// TIA Portal project "Konzept_zur_Überwachung_der_Feuchtigkeit_des_Getriebeöls" (V18)

(* hardware
DEVICE "Haupt_Station"  TP2200 Comfort
   slot 0: "Haupt_Station"  TP2200 Comfort  6AV2 124-0XC02-0AX0  17.0.0.0
   slot 1: "HMI_RT"  TP2200 Comfort  6AV2 124-0XC02-0AX0  17.0.0.0
   slot 5: "Haupt_Station.IE_CP_2"  PROFINET Interface  17.0.0.0
      slot 1: "PROFINET Schnittstelle_1"  PROFINET Interface
         slot 1: "Port_1"  Port
         slot 2: "Port_2"  Port
   slot 6: "Haupt_Station.IE_CP_1"  PROFINET Interface  17.0.0.0
      slot 1: "PROFINET Schnittstelle_GBit"  PROFINET Interface
         slot 1: "Port_1"  Port
   slot 7: "Haupt_Station.MPI/DP_CP_1"  MPI/DP Interface  17.0.0.0
DEVICE "S7-1500/ET200MP-Station_1"  S7-1500 station
   slot 0: "Profilschiene_0"  Rack  6ES7 590-1***0-0AA0
   slot 1: "1513"  CPU 1513-1 PN  6ES7 513-1AM03-0AB0  V3.0
      slot 3: "CPU-Display_1"  6ES7591-1AA00-0AA0
      slot 32768: "PROFINET-Schnittstelle_1"  X1
         slot 32769: "Port_1"  X1 P1
         slot 32770: "Port_2"  X1 P2
      slot 34817: "Virtual CP interface port_1"  Virtual CP interface port  Virtual CP interface port
   slot 2: "DI 16x24VDC / DQ 16x24VDC/0.5A BA_1"  DI 16x24VDC/DQ 16x24VDC/0.5A BA  6ES7 523-1BL00-0AA0  V1.1
   slot 3: "AI 8xU/I/R/RTD BA_1"  AI 8xU/I/R/RTD BA  6ES7 531-7QF00-0AB0  V1.0
DEVICE "S7-300/ET200M-Station_1"  S7-300 station
   slot 0: "Profilschiene_0"  Rail  6ES7 390-1***0-0AA0
   slot 1: "PS 307 10A_1"  PS 307 10A  6ES7 307-1KA02-0AA0
   slot 2: "313C"  CPU 313C-2 DP  6ES7 313-6CG04-0AB0  V3.3
      slot 0: "MPI-Schnittstelle_1"  MPI
      slot 1: "DP-Schnittstelle_1"  DP
      slot 2: "DI 16/DO 16_1"  DI16/DO16
      slot 4: "Zählen_1"  Counter
   slot 4: "AI 8x13BIT_1"  AI8x13Bit  6ES7 331-1KF02-0AB0
*)

// ===== PLC "1513"  CPU 1513-1 PN =====

VAR_GLOBAL   // PLC tag table "Standard-Variablentabelle"
   "LDH_Temp_1(1)" AT %IW34 : Int;
   "LDH_Feucht_1(1)" AT %IW36 : Int;
   "LDH_Temp_2(1)" AT %IW38 : Int;
   "LDH_Feucht_2(1)" AT %IW40 : Int;
   "Gill_Fine(1)" AT %IW42 : Int;
   "Gill_Coarse(1)" AT %IW44 : Int;
   "Gill_Water(1)" AT %IW46 : Int;
   "Gill_Fehler(1)" AT %IW48 : Int;
   "Rote_Lampe(1)" AT %Q0.0 : Bool;
   "Orange_Lampe(1)" AT %Q0.1 : Bool;
   "Grüne_Lampe_2(1)" AT %Q0.2 : Bool;
   "Abschalten_M(1)" AT %Q0.3 : Bool;
   "Quittierung(1)" AT %I0.0 : Bool;
END_VAR

DATA_BLOCK "Rt_Zyklus_DB"   // DB1
{ S7_Optimized_Access := 'TRUE' }
VERSION : 0.1
// stored: InstanceOfName Rt_Zyklus
"Rt_Zyklus"
BEGIN
END_DATA_BLOCK

DATA_BLOCK "LDH100_DB_1"   // DB2
{ S7_Optimized_Access := 'TRUE' }
VERSION : 0.1
// stored: InstanceOfName LDH100
"LDH100"
BEGIN
END_DATA_BLOCK

DATA_BLOCK "LDH100_DB_2"   // DB3
{ S7_Optimized_Access := 'TRUE' }
VERSION : 0.1
// stored: InstanceOfName LDH100
"LDH100"
BEGIN
END_DATA_BLOCK

DATA_BLOCK "GILL4212_DB"   // DB4
{ S7_Optimized_Access := 'TRUE' }
VERSION : 0.1
// stored: InstanceOfName GILL4212
"GILL4212"
BEGIN
END_DATA_BLOCK

DATA_BLOCK "HMI"   // DB5
{ S7_Optimized_Access := 'TRUE' }
VERSION : 0.1
   VAR
      Quittieren1500 : Bool;
   END_VAR
BEGIN
END_DATA_BLOCK

FUNCTION_BLOCK "LDH100"   // FB1, SCL
{ S7_Optimized_Access := 'TRUE' }
VERSION : 0.1
   VAR_INPUT
      AI_Temp_RAW : Int;
      cycleTime_ms : Real;
      AI_Hum_RAW : Int;
      Quittieren : Bool;
   END_VAR
   VAR_OUTPUT
      Temp_filt : Real;
      Temp_real : Real;
      Hum_filt : Real;
      Hum_real : Real;
      Warnung : Bool;
      Alarm_Temp : Bool;
      Alarm_Hum : Bool;
      OK : Bool;
      SensorError_Temp : Bool;
      SensorError_Hum : Bool;
      SensorDefekt : Bool;
      Strom_Temp_mA : Real;
      Strom_Hum_mA : Real;
   END_VAR
   VAR
      Alarm_Temp_Intern : Bool;
      TempGrenze_Alarm : Real := 0.0;
      HumGrenze_Alarm : Real := 0.0;
      Alarm_Hum_Intern : Bool;
      intervall_temp : Real;
      intervall_hum : Real;
      TON_temp : TON_TIME;
      TON_Hum : TON_TIME;
      RawTol : Int;
      RawMin : Int;
      RawMax : Int;
   END_VAR
   VAR_TEMP
      Norm_Temp : Real;
      alpha_pt1 : Real;
      Norm_Hum : Real;
   END_VAR
   VAR CONSTANT
      T_PT1_ms : Real := 565.0;
   END_VAR
BEGIN
   // -2) Rohwert-Toleranz (±0,2 mA auf 4–>20 mA = -346–>27648)
   #RawTol := REAL_TO_INT((0.2 / 16.0) * 27648.0);
   #RawMin := - #RawTol;
   #RawMax := 27648 + #RawTol;

   // -1) Strom in mA berechnen
   #Strom_Temp_mA := (INT_TO_REAL(#AI_Temp_RAW) / 27648.0) * 16.0 + 4.0;
   #Strom_Hum_mA := (INT_TO_REAL(#AI_Hum_RAW) / 27648.0) * 16.0 + 4.0;

   // 0) Sensor-Error prüfen auf Rohwerte
   #SensorError_Temp := (#AI_Temp_RAW < #RawMin) OR (#AI_Temp_RAW > #RawMax);
   #SensorError_Hum := (#AI_Hum_RAW < #RawMin) OR (#AI_Hum_RAW > #RawMax);

   // 1) Skalierung in reale Werte
   #Temp_real := (INT_TO_REAL(#AI_Temp_RAW) / 27648.0) * 140.0 - 20.0;  // -20°C ... +120°C
   #Hum_real := (INT_TO_REAL(#AI_Hum_RAW) / 27648.0) * 100.0;         // 0% ... 100%

   // 2) Filter-Koeffizient berechnen (für τ = 565 ms → 90 % nach 1.3 s)
   #alpha_pt1 := #cycleTime_ms / (#T_PT1_ms + #cycleTime_ms);

   // 3) PT1-Glättung
   #Temp_filt := #Temp_filt + #alpha_pt1 * (#Temp_real - #Temp_filt);
   #Hum_filt := #Hum_filt + #alpha_pt1 * (#Hum_real - #Hum_filt);

   // 4) Alarm-Logik mit IEC-Timer (TON)
   // → nur auslösen, wenn Filterwert 1.3 s lang über Grenzwert liegt
   #TON_temp(IN := (#Temp_filt >= #TempGrenze_Alarm),
             PT := T#1300ms);
   #TON_Hum(IN := (#Hum_filt >= #HumGrenze_Alarm),
            PT := T#1300ms);

   IF #TON_temp.Q THEN
       #Alarm_Temp := TRUE;
   ELSIF #Quittieren AND (#Temp_filt < #TempGrenze_Alarm) THEN
       #Alarm_Temp := FALSE;
   END_IF;

   IF #TON_Hum.Q THEN
       #Alarm_Hum := TRUE;
   ELSIF #Quittieren AND (#Hum_filt < #HumGrenze_Alarm) THEN
       #Alarm_Hum := FALSE;
   END_IF;

   // 5) Warnung (Echtwerte, keine Filterung nötig)
   #Warnung := (#Temp_real >= (#TempGrenze_Alarm - #intervall_temp)) OR
   (#Hum_real >= (#HumGrenze_Alarm - #intervall_hum));

   // 6) OK-Status
   #OK := NOT #Alarm_Temp AND NOT #Alarm_Hum;
END_FUNCTION_BLOCK

FUNCTION_BLOCK "GILL4212"   // FB2, SCL
{ S7_Optimized_Access := 'TRUE' }
VERSION : 0.1
   VAR_INPUT
      AI_Fine_RAW : Int;
      AI_Coarse_RAW : Int;
      AI_Water_RAW : Int;
      Quittieren : Bool;
   END_VAR
   VAR_OUTPUT
      SensorError_Coarse : Bool;
      SensorError_Water : Bool;
      SensorError_Fine : Bool;
      Fine_percent : Real;
      Coarse_percent : Real;
      Water_percent : Real;
      Alarm_Wear : Bool;
      Alarm_Water : Bool;
      Warnung : Bool;
      OK : Bool;
   END_VAR
   VAR
      TON_Wear : TON_TIME;
      TON_Water : TON_TIME;
      Alarm_Wear_Intern : Bool;
      Alarm_Water_Intern : Bool;
      RawTol : Int;
      RawMin : Int;
      RawMax : Int;
   END_VAR
   VAR CONSTANT
      Wear_Alarm_Limit : Real := 70.0;
      Water_Alarm_Limit : Real := 60.0;
   END_VAR
BEGIN
   // -1) Toleranzbereich in Rohwert berechnen (±0.2 mA)
   #RawTol := REAL_TO_INT((0.2 / 16.0) * 27648.0);
   #RawMin := - #RawTol;
   #RawMax := 27648 + #RawTol;

   // 0) Rohwert auf Gültigkeit prüfen (Toleranz)
   #SensorError_Fine := (#AI_Fine_RAW < #RawMin) OR (#AI_Fine_RAW > #RawMax);
   #SensorError_Coarse := (#AI_Coarse_RAW < #RawMin) OR (#AI_Coarse_RAW > #RawMax);
   #SensorError_Water := (#AI_Water_RAW < #RawMin) OR (#AI_Water_RAW > #RawMax);

   // 1) Skalierung 4–20 mA → 0–100 %
   #Fine_percent := (INT_TO_REAL(#AI_Fine_RAW) / 27648.0) * 100.0;
   #Coarse_percent := (INT_TO_REAL(#AI_Coarse_RAW) / 27648.0) * 100.0;
   #Water_percent := (INT_TO_REAL(#AI_Water_RAW) / 27648.0) * 100.0;

   // 2) Alarmverzögerung (1,3 Sekunden) mit TON
   #TON_Wear(IN := (#Fine_percent >= #Wear_Alarm_Limit) OR (#Coarse_percent >= #Wear_Alarm_Limit), PT := T#1300ms);
   #TON_Water(IN := (#Water_percent >= #Water_Alarm_Limit), PT := T#1300ms);

   // 3) Alarm setzen nach Ablauf der Verzögerung
   IF #TON_Wear.Q THEN
       #Alarm_Wear_Intern := TRUE;
   END_IF;
   IF #TON_Water.Q THEN
       #Alarm_Water_Intern := TRUE;
   END_IF;

   // 4) Quittierung (nur wenn alle Werte unterhalb der Limits)
   IF #Quittieren AND #Fine_percent < #Wear_Alarm_Limit AND #Coarse_percent < #Wear_Alarm_Limit THEN
       #Alarm_Wear_Intern := FALSE;
   END_IF;
   IF #Quittieren AND #Water_percent < #Water_Alarm_Limit THEN
       #Alarm_Water_Intern := FALSE;
   END_IF;

   // 5) Ausgänge setzen
   #Alarm_Wear := #Alarm_Wear_Intern;
   #Alarm_Water := #Alarm_Water_Intern;

   // 6) Warnung (Vorwarnbereich ohne Verzögerung)
   #Warnung :=
   (#Fine_percent >= #Wear_Alarm_Limit - 20.0) OR
   (#Coarse_percent >= #Wear_Alarm_Limit - 20.0) OR
   (#Water_percent >= #Water_Alarm_Limit - 20.0);

   // 7) OK-Status
   #OK := NOT #Alarm_Wear AND NOT #Alarm_Water;
END_FUNCTION_BLOCK

FUNCTION_BLOCK "Rt_Zyklus"   // FB3, SCL
{ S7_Optimized_Access := 'TRUE' }
VERSION : 0.1
   VAR_INPUT
      Enable : Bool := True;
      Reset : Bool;
   END_VAR
   VAR_OUTPUT
      Cycle_ms : LReal;
      Min_ms : LReal;
      Max_ms : LReal;
      Error : Bool;
      Status : Int;
   END_VAR
   VAR
      Last_ns : LTime;
      Min_ns : LTime;
      Max_ns : LTime;
      ResetOld : Bool;
   END_VAR
BEGIN

   IF #Enable THEN

       // --- 1) Letzte Zykluszeit holen -----------------------------
       #Status := RT_INFO(
                          MODE := 25,          // MODE 25 = letzte Zykluszeit
                          OB := 0,
                          INFO := #Last_ns     // LTIME (Nanosekunden)
       );

   // Fehlerbehandlung -------------------------------------------
   #Error:= (#Status <> 0); // 0 = OK, alles andere = Fehler


       IF NOT #Error THEN

           // --- 2) Umrechnen in Millisekunden ----------------------
           #Cycle_ms := LINT_TO_LREAL(#Last_ns) / 1_000_000.0;

           // --- 3) Min/Max bilden ---------------------------------
           IF #Last_ns < #Min_ns THEN
               #Min_ns := #Last_ns;
           END_IF;

           IF #Last_ns > #Max_ns THEN
               #Max_ns := #Last_ns;
           END_IF;

           // --- 4) Reset per Flanke --------------------------------
           IF #Reset AND NOT #ResetOld THEN      // positive Flanke
               #Min_ns := #Last_ns;
               #Max_ns := #Last_ns;
           END_IF;

           // --- 5) Ausgänge aktualisieren --------------------------
           #Min_ms := LINT_TO_LREAL(#Min_ns) / 1_000_000.0;
           #Max_ms := LINT_TO_LREAL(#Max_ns) / 1_000_000.0;
       END_IF;

       // Flankenerkennung speicher­n
       #ResetOld := #Reset;

   ELSE
       // Messung deaktiviert → keine neuen Werte bilden
       #Error := FALSE;
       #Status := 0;
   END_IF;
END_FUNCTION_BLOCK

FUNCTION "Ampel_Logik" : Void   // FC1, SCL
{ S7_Optimized_Access := 'TRUE' }
VERSION : 0.1
   VAR_INPUT
      LDH1_Alarm_Hum : Bool;   // Alarm von LDH1 (Feuchte)
      LDH1_Alarm_Temp : Bool;   // Alarm von LDH1 (Temperatur)
      LDH2_Alarm_Hum : Bool;   // Alarm von LDH2 (Feuchte)
      LDH2_Alarm_Temp : Bool;   // Alarm von LDH2 (Temperatur)
      GILL_Alarm_Wear : Bool;   // Alarm vom GILL-Sensor (Verschleiß)
      GILL_Alarm_Water : Bool;   // Alarm vom GILL-Sensor (Wasser)
      LDH1_Warnung : Bool;   // Warnung LDH100_1
      LDH2_Warnung : Bool;   // Warnung LDH100_1
      GILL_Warnung : Bool;   // Warnung Verschleiss
   END_VAR
   VAR_OUTPUT
      LAMP_ROT : Bool;
      LAMP_ORANGE : Bool;
      LAMP_GRUEN : Bool;
   END_VAR
   VAR CONSTANT
      TempWarnMin : Real := 80.0;
      HumWarnMin : Real := 40.0;
      WearWarnMin : Real := 70.0;
      WaterWarnMin : Real := 50.0;
      HumAlarmLimit : Real := 100.0;
      TempAlarmLimit : Real := 60.0;
      WearAlarmLimit : Real := 80.0;
      WaterAlarmLimit : Real := 60.0;
   END_VAR
BEGIN
   // 1) ROT: mindestens ein Alarm-Flag aktiv
   IF #LDH1_Alarm_Hum OR #LDH1_Alarm_Temp OR
       #LDH2_Alarm_Hum OR #LDH2_Alarm_Temp OR
       #GILL_Alarm_Wear OR #GILL_Alarm_Water THEN

       #LAMP_ROT := TRUE;
       #LAMP_ORANGE := FALSE;
       #LAMP_GRUEN := FALSE;

       // 2) ORANGE: mindestens ein Wert im Warnbereich
       // 2) ORANGE: mindestens ein Warn-Flag aktiv
   ELSIF #LDH1_Warnung OR #LDH2_Warnung OR #GILL_Warnung THEN

       #LAMP_ROT := FALSE;
       #LAMP_ORANGE := TRUE;
       #LAMP_GRUEN := FALSE;

       // 3) GRÜN: alle Werte unter Warnschwelle
   ELSE
       #LAMP_ROT := FALSE;
       #LAMP_ORANGE := FALSE;
       #LAMP_GRUEN := TRUE;
   END_IF;
END_FUNCTION

ORGANIZATION_BLOCK "Main"   // OB1, LAD, ProgramCycle
TITLE = "Main Program Sweep (Cycle)"
{ S7_Optimized_Access := 'TRUE' }
VERSION : 0.1
   VAR_INPUT
      Initial_Call : Bool;   // Initial call of this OB
      Remanence : Bool;   // =True, if remanent data are available
   END_VAR
BEGIN

REGION Network 1
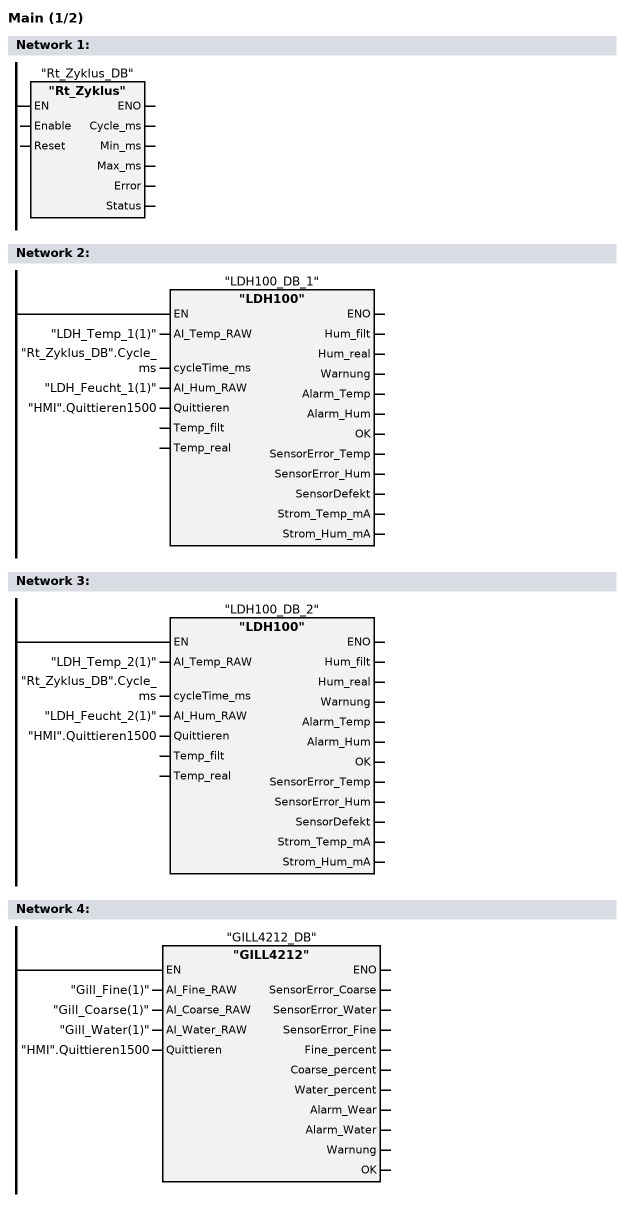
   RUNG wire#powerrail
      "Rt_Zyklus_DB"(Enable :=, Reset :=, Cycle_ms =>, Min_ms =>, Max_ms =>, Error =>, Status =>)
   END_RUNG
   // the same network as SCL:
   "Rt_Zyklus_DB"();   // "Rt_Zyklus"
END_REGION

REGION Network 2
   RUNG wire#powerrail
      "LDH100_DB_1"(AI_Temp_RAW := "LDH_Temp_1(1)", cycleTime_ms := "Rt_Zyklus_DB".Cycle_ms, AI_Hum_RAW := "LDH_Feucht_1(1)", Quittieren := "HMI".Quittieren1500, Temp_filt :=, Temp_real :=, Hum_filt =>, Hum_real =>, Warnung =>, Alarm_Temp =>, Alarm_Hum =>, OK =>, SensorError_Temp =>, SensorError_Hum =>, SensorDefekt =>, Strom_Temp_mA =>, Strom_Hum_mA =>)
   END_RUNG
   // the same network as SCL:
   "LDH100_DB_1"(AI_Temp_RAW := "LDH_Temp_1(1)",   // "LDH100"
                 cycleTime_ms := "Rt_Zyklus_DB".Cycle_ms,
                 AI_Hum_RAW := "LDH_Feucht_1(1)",
                 Quittieren := "HMI".Quittieren1500);
END_REGION

REGION Network 3
   RUNG wire#powerrail
      "LDH100_DB_2"(AI_Temp_RAW := "LDH_Temp_2(1)", cycleTime_ms := "Rt_Zyklus_DB".Cycle_ms, AI_Hum_RAW := "LDH_Feucht_2(1)", Quittieren := "HMI".Quittieren1500, Temp_filt :=, Temp_real :=, Hum_filt =>, Hum_real =>, Warnung =>, Alarm_Temp =>, Alarm_Hum =>, OK =>, SensorError_Temp =>, SensorError_Hum =>, SensorDefekt =>, Strom_Temp_mA =>, Strom_Hum_mA =>)
   END_RUNG
   // the same network as SCL:
   "LDH100_DB_2"(AI_Temp_RAW := "LDH_Temp_2(1)",   // "LDH100"
                 cycleTime_ms := "Rt_Zyklus_DB".Cycle_ms,
                 AI_Hum_RAW := "LDH_Feucht_2(1)",
                 Quittieren := "HMI".Quittieren1500);
END_REGION

REGION Network 4
   RUNG wire#powerrail
      "GILL4212_DB"(AI_Fine_RAW := "Gill_Fine(1)", AI_Coarse_RAW := "Gill_Coarse(1)", AI_Water_RAW := "Gill_Water(1)", Quittieren := "HMI".Quittieren1500, SensorError_Coarse =>, SensorError_Water =>, SensorError_Fine =>, Fine_percent =>, Coarse_percent =>, Water_percent =>, Alarm_Wear =>, Alarm_Water =>, Warnung =>, OK =>)
   END_RUNG
   // the same network as SCL:
   "GILL4212_DB"(AI_Fine_RAW := "Gill_Fine(1)",   // "GILL4212"
                 AI_Coarse_RAW := "Gill_Coarse(1)",
                 AI_Water_RAW := "Gill_Water(1)",
                 Quittieren := "HMI".Quittieren1500);
END_REGION

REGION Network 5
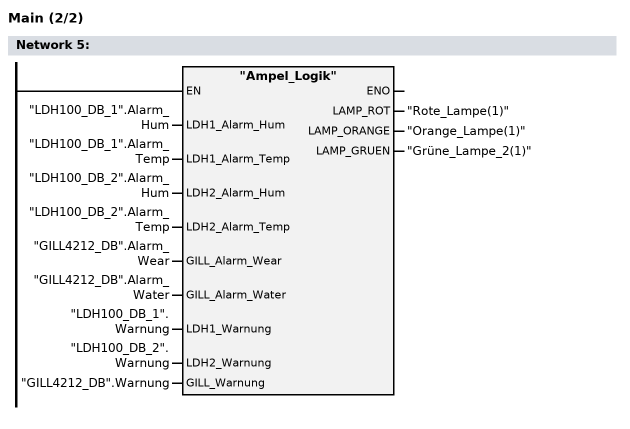
   RUNG wire#powerrail
      "Ampel_Logik"(LDH1_Alarm_Hum := "LDH100_DB_1".Alarm_Hum, LDH1_Alarm_Temp := "LDH100_DB_1".Alarm_Temp, LDH2_Alarm_Hum := "LDH100_DB_2".Alarm_Hum, LDH2_Alarm_Temp := "LDH100_DB_2".Alarm_Temp, GILL_Alarm_Wear := "GILL4212_DB".Alarm_Wear, GILL_Alarm_Water := "GILL4212_DB".Alarm_Water, LDH1_Warnung := "LDH100_DB_1".Warnung, LDH2_Warnung := "LDH100_DB_2".Warnung, GILL_Warnung := "GILL4212_DB".Warnung, LAMP_ROT => "Rote_Lampe(1)", LAMP_ORANGE => "Orange_Lampe(1)", LAMP_GRUEN => "Grüne_Lampe_2(1)")
   END_RUNG
   // the same network as SCL:
   "Ampel_Logik"(LDH1_Alarm_Hum := "LDH100_DB_1".Alarm_Hum,
                 LDH1_Alarm_Temp := "LDH100_DB_1".Alarm_Temp,
                 LDH2_Alarm_Hum := "LDH100_DB_2".Alarm_Hum,
                 LDH2_Alarm_Temp := "LDH100_DB_2".Alarm_Temp,
                 GILL_Alarm_Wear := "GILL4212_DB".Alarm_Wear,
                 GILL_Alarm_Water := "GILL4212_DB".Alarm_Water,
                 LDH1_Warnung := "LDH100_DB_1".Warnung,
                 LDH2_Warnung := "LDH100_DB_2".Warnung,
                 GILL_Warnung := "GILL4212_DB".Warnung,
                 LAMP_ROT => "Rote_Lampe(1)",
                 LAMP_ORANGE => "Orange_Lampe(1)",
                 LAMP_GRUEN => "Grüne_Lampe_2(1)");
END_REGION
END_ORGANIZATION_BLOCK

// ===== PLC "313C"  CPU 313C-2 DP =====

VAR_GLOBAL   // PLC tag table "Standard-Variablentabelle"
   "LDH_Temp_1" AT %IW272 : Int;
   "LDH_Feucht_1" AT %IW274 : Int;
   "LDH_Temp_2" AT %IW276 : Int;
   "LDH_Feucht_2" AT %IW278 : Int;
   "Gill_Fine" AT %IW280 : Int;
   "Gill_Coarse" AT %IW282 : Int;
   "Gill_Water" AT %IW284 : Int;
   "Gill_Fehler" AT %IW286 : Int;
   "Rote_Lampe" AT %I124.0 : Bool;
   "Orange_Lampe" AT %I124.1 : Bool;
   "Grüne_Lampe_2" AT %I124.2 : Bool;
   "Abschalten_M" AT %I124.3 : Bool;
END_VAR

VAR_GLOBAL   // PLC tag table "Merker_B"
   "B1" AT %M0.0 : Bool;
   "B2" AT %M0.1 : Bool;
   "B3" AT %M0.2 : Bool;
   "B4" AT %M0.3 : Bool;
   "B5" AT %M0.4 : Bool;
   "Re1" AT %MD1 : Real;
   "Re2" AT %MD2 : Real;
   "Re3" AT %MD3 : Real;
   "Re4" AT %MD4 : Real;
   "B7" AT %M0.6 : Bool;
   "B6" AT %M0.5 : Bool;
   "Re5" AT %MD5 : Real;
   "Re6" AT %MD6 : Real;
END_VAR

DATA_BLOCK "LDH100_DB_1"   // DB1
{ S7_Optimized_Access := 'FALSE' }
VERSION : 0.1
// stored: InstanceOfName LDH100
"LDH100"
BEGIN
   TempGrenze_Alarm := 60.0;
   HumGrenze_Alarm := 90.0;
   intervall_temp := 10.0;
   intervall_hum := 20.0;
END_DATA_BLOCK

DATA_BLOCK "LDH100_DB_2"   // DB2
{ S7_Optimized_Access := 'FALSE' }
VERSION : 0.1
// stored: InstanceOfName LDH100
"LDH100"
BEGIN
END_DATA_BLOCK

DATA_BLOCK "GILL4212_DB"   // DB3
{ S7_Optimized_Access := 'FALSE' }
VERSION : 0.1
// stored: InstanceOfName GILL4212
"GILL4212"
BEGIN
END_DATA_BLOCK

DATA_BLOCK "HMI_313"   // DB4
{ S7_Optimized_Access := 'FALSE' }
VERSION : 0.1
   VAR
      Quittieren313 : Bool;
   END_VAR
BEGIN
END_DATA_BLOCK

FUNCTION_BLOCK "LDH100"   // FB1, SCL
{ S7_Optimized_Access := 'FALSE' }
VERSION : 0.1
   VAR_INPUT
      AI_Temp_RAW : Int;
      cycleTime_ms : Int;
      AI_Hum_RAW : Int;
      Quittieren : Bool;
   END_VAR
   VAR_OUTPUT
      Temp_filt : Real;
      Hum_filt : Real;
      Temp_real : Real;
      Hum_real : Real;
      Warnung : Bool;
      OK : Bool;
      SensorError_Temp : Bool;
      SensorError_Hum : Bool;
      SensorDefekt : Bool;
      Strom_Hum_mA : Real;
      Strom_Temp_mA : Real;
      Alarm_Temp : Bool;
      Alarm_Hum : Bool;
   END_VAR
   VAR
      Alarm_Temp_Intern : Bool;
      TempGrenze_Alarm : Real := 0.0;
      HumGrenze_Alarm : Real := 0.0;
      Alarm_Hum_Intern : Bool;
      intervall_temp : Real;
      intervall_hum : Real;
      RawTol : Int;
      RawMin : Int;
      cycleTime_s : Real;
      TON_temp : TON;
      TON_Hum : TON;
      RawMax : Int;
   END_VAR
   VAR_TEMP
      Norm_Temp : Real;
      alpha_pt1 : Real;
      Norm_Hum : Real;
   END_VAR
   VAR CONSTANT
      T_PT1_ms : Real := 565.0;
      tSensorDelay : Time := T#1300ms;
   END_VAR
BEGIN
   // -2) Rohwert-Toleranz (±0,2 mA auf 4–>20 mA = -346–>27648)
   #RawTol := REAL_TO_INT((0.2 / 16.0) * 27648.0);  
   #RawMin := -#RawTol;                                     
   #RawMax := 27648 + #RawTol;

   // -1) Strom in mA berechnen
   #Strom_Temp_mA := (INT_TO_REAL(#AI_Temp_RAW) / 27648.0) * 16.0 + 4.0;
   #Strom_Hum_mA := (INT_TO_REAL(#AI_Hum_RAW) / 27648.0) * 16.0 + 4.0;

   // 0) Sensor-Error prüfen auf Rohwerte
   #SensorError_Temp := (#AI_Temp_RAW < #RawMin) OR (#AI_Temp_RAW > #RawMax);
   #SensorError_Hum := (#AI_Hum_RAW < #RawMin) OR (#AI_Hum_RAW > #RawMax);

   // 1) Skalierung in reale Werte
   #Temp_real := (INT_TO_REAL(#AI_Temp_RAW) / 27648.0) * 140.0 - 20.0;  // -20°C ... +120°C
   #Hum_real := (INT_TO_REAL(#AI_Hum_RAW) / 27648.0) * 100.0;         // 0% ... 100%

   // 2) Filter-Koeffizient berechnen (für τ = 565 ms → 90 % nach 1.3 s)
   #alpha_pt1 := INT_TO_REAL(#cycleTime_ms) / (#T_PT1_ms + INT_TO_REAL(#cycleTime_ms));

   // 3) PT1-Glättung
   #Temp_filt := #Temp_filt + #alpha_pt1 * (#Temp_real - #Temp_filt);
   #Hum_filt := #Hum_filt + #alpha_pt1 * (#Hum_real - #Hum_filt);

   // 4) Alarm-Logik mit IEC-Timer (TON)
   // → nur auslösen, wenn Filterwert 1.3 s lang über Grenzwert liegt
   #TON_temp(IN := (#Temp_filt >= #TempGrenze_Alarm), PT := T#1300ms);
   #TON_Hum(IN  := (#Hum_filt  >= #HumGrenze_Alarm),  PT := T#1300ms);

   IF #TON_temp.Q THEN
       #Alarm_Temp := TRUE;
   ELSIF #Quittieren AND (#Temp_filt < #TempGrenze_Alarm) THEN
       #Alarm_Temp := FALSE;
   END_IF;

   IF #TON_Hum.Q THEN
       #Alarm_Hum := TRUE;
   ELSIF #Quittieren AND (#Hum_filt < #HumGrenze_Alarm) THEN
       #Alarm_Hum := FALSE;
   END_IF;

   // 5) Warnung (Echtwerte, keine Filterung nötig)
   #Warnung := (#Temp_real >= (#TempGrenze_Alarm - #intervall_temp)) OR
   (#Hum_real >= (#HumGrenze_Alarm - #intervall_hum));

   // 6) OK-Status
   #OK := NOT #Alarm_Temp AND NOT #Alarm_Hum;
END_FUNCTION_BLOCK

FUNCTION_BLOCK "GILL4212"   // FB2, SCL
{ S7_Optimized_Access := 'FALSE' }
VERSION : 0.1
   VAR_INPUT
      AI_Fine_RAW : Int;
      AI_Coarse_RAW : Int;
      AI_Water_RAW : Int;
      Quittieren : Bool;
   END_VAR
   VAR_OUTPUT
      Fine_percent : Real;
      Coarse_percent : Real;
      Water_percent : Real;
      Alarm_Wear : Bool;
      Alarm_Water : Bool;
      Warnung : Bool;
      SensorError_Coarse : Bool;
      SensorError_Water : Bool;
      SensorError_Fine : Bool;
      OK : Bool;
   END_VAR
   VAR
      Alarm_Wear_Intern : Bool;
      Alarm_Water_Intern : Bool;
      RawTol : Int;
      RawMin : Int;
      TON_Wear : TON;
      TON_Water : TON;
      RawMax : Int;
   END_VAR
   VAR CONSTANT
      Wear_Alarm_Limit : Real := 70.0;
      Water_Alarm_Limit : Real := 60.0;
   END_VAR
BEGIN
   // -1) Toleranzbereich in Rohwert berechnen (±0.2 mA)
   #RawTol := REAL_TO_INT((0.2 / 16.0) * 27648.0);
   #RawMin := - #RawTol;
   #RawMax := 27648 + #RawTol;

   // 0) Rohwert auf Gültigkeit prüfen (Toleranz)
   #SensorError_Fine := (#AI_Fine_RAW < #RawMin) OR (#AI_Fine_RAW > #RawMax);
   #SensorError_Coarse := (#AI_Coarse_RAW < #RawMin) OR (#AI_Coarse_RAW > #RawMax);
   #SensorError_Water := (#AI_Water_RAW < #RawMin) OR (#AI_Water_RAW > #RawMax);

   // 1) Skalierung 4–20 mA → 0–100 %
   #Fine_percent := (INT_TO_REAL(#AI_Fine_RAW) / 27648.0) * 100.0;
   #Coarse_percent := (INT_TO_REAL(#AI_Coarse_RAW) / 27648.0) * 100.0;
   #Water_percent := (INT_TO_REAL(#AI_Water_RAW) / 27648.0) * 100.0;

   // 2) Alarmverzögerung (1,3 Sekunden) mit TON
   #TON_Wear(IN := (#Fine_percent >= #Wear_Alarm_Limit) OR (#Coarse_percent >= #Wear_Alarm_Limit), PT := T#1300ms);
   #TON_Water(IN := (#Water_percent >= #Water_Alarm_Limit), PT := T#1300ms);

   // 3) Alarm setzen nach Ablauf der Verzögerung
   IF #TON_Wear.Q THEN
       #Alarm_Wear_Intern := TRUE;
   END_IF;
   IF #TON_Water.Q THEN
       #Alarm_Water_Intern := TRUE;
   END_IF;

   // 4) Quittierung (nur wenn alle Werte unterhalb der Limits)
   IF #Quittieren AND #Fine_percent < #Wear_Alarm_Limit AND #Coarse_percent < #Wear_Alarm_Limit THEN
       #Alarm_Wear_Intern := FALSE;
   END_IF;
   IF #Quittieren AND #Water_percent < #Water_Alarm_Limit THEN
       #Alarm_Water_Intern := FALSE;
   END_IF;

   // 5) Ausgänge setzen
   #Alarm_Wear := #Alarm_Wear_Intern;
   #Alarm_Water := #Alarm_Water_Intern;

   // 6) Warnung (Vorwarnbereich ohne Verzögerung)
   #Warnung :=
   (#Fine_percent >= #Wear_Alarm_Limit - 20.0) OR
   (#Coarse_percent >= #Wear_Alarm_Limit - 20.0) OR
   (#Water_percent >= #Water_Alarm_Limit - 20.0);

   // 7) OK-Status
   #OK := NOT #Alarm_Wear AND NOT #Alarm_Water;
END_FUNCTION_BLOCK

FUNCTION "Ampel_Logik" : Void   // FC1, SCL
{ S7_Optimized_Access := 'FALSE' }
VERSION : 0.1
   VAR_INPUT
      LDH1_Alarm_Hum : Bool;   // Alarm von LDH1 (Feuchte)
      LDH1_Alarm_Temp : Bool;   // Alarm von LDH1 (Temperatur)
      LDH2_Alarm_Hum : Bool;   // Alarm von LDH2 (Feuchte)
      LDH2_Alarm_Temp : Bool;   // Alarm von LDH2 (Temperatur)
      GILL_Alarm_Wear : Bool;   // Alarm vom GILL-Sensor (Verschleiß)
      GILL_Alarm_Water : Bool;   // Alarm vom GILL-Sensor (Wasser)
      LDH1_Warnung : Bool;   // Warnung LDH100_1
      LDH2_Warnung : Bool;   // Warnung LDH100_1
      GILL_Warnung : Bool;   // Warnung Verschleiss
   END_VAR
   VAR_OUTPUT
      LAMP_ROT : Bool;
      LAMP_ORANGE : Bool;
      LAMP_GRUEN : Bool;
   END_VAR
   VAR CONSTANT
      TempWarnMin : Real := 80.0;
      HumWarnMin : Real := 40.0;
      WearWarnMin : Real := 70.0;
      WaterWarnMin : Real := 50.0;
      HumAlarmLimit : Real := 100.0;
      TempAlarmLimit : Real := 60.0;
      WearAlarmLimit : Real := 80.0;
      WaterAlarmLimit : Real := 60.0;
   END_VAR
BEGIN
   // 1) ROT: mindestens ein Alarm-Flag aktiv
   IF #LDH1_Alarm_Hum OR #LDH1_Alarm_Temp OR
       #LDH2_Alarm_Hum OR #LDH2_Alarm_Temp OR
       #GILL_Alarm_Wear OR #GILL_Alarm_Water THEN

       #LAMP_ROT := TRUE;
       #LAMP_ORANGE := FALSE;
       #LAMP_GRUEN := FALSE;

       // 2) ORANGE: mindestens ein Wert im Warnbereich
       // 2) ORANGE: mindestens ein Warn-Flag aktiv
   ELSIF #LDH1_Warnung OR #LDH2_Warnung OR #GILL_Warnung THEN

       #LAMP_ROT := FALSE;
       #LAMP_ORANGE := TRUE;
       #LAMP_GRUEN := FALSE;

       // 3) GRÜN: alle Werte unter Warnschwelle
   ELSE
       #LAMP_ROT := FALSE;
       #LAMP_ORANGE := FALSE;
       #LAMP_GRUEN := TRUE;
   END_IF;
END_FUNCTION

ORGANIZATION_BLOCK "Main"   // OB1, LAD
TITLE = "Main Program Sweep (Cycle)"
{ S7_Optimized_Access := 'FALSE' }
VERSION : 0.1
   VAR_TEMP
      OB1_EV_CLASS : Byte;   // Bits 0-3 = 1 (Coming event), Bits 4-7 = 1 (Event class 1)
      OB1_SCAN_1 : Byte;   // 1 (Cold restart scan 1 of OB 1), 3 (Scan 2-n of OB 1)
      OB1_PRIORITY : Byte;   // Priority of OB Execution
      OB1_OB_NUMBR : Byte;   // 1 (Organization block 1, OB1)
      OB1_RESERVED_1 : Byte;   // Reserved for system
      OB1_RESERVED_2 : Byte;   // Reserved for system
      OB1_PREV_CYCLE : Int;   // Cycle time of previous OB1 scan (milliseconds)
      OB1_MIN_CYCLE : Int;   // Minimum cycle time of OB1 (milliseconds)
      OB1_MAX_CYCLE : Int;   // Maximum cycle time of OB1 (milliseconds)
      OB1_DATE_TIME : Date_And_Time;   // Date and time OB1 started
   END_VAR
BEGIN

REGION Network 1
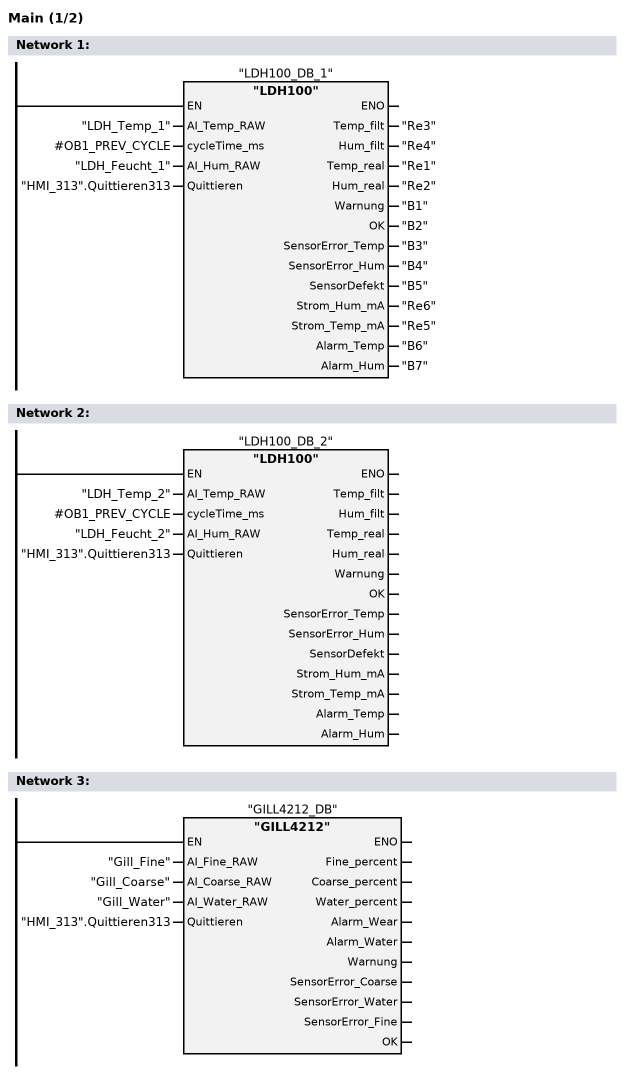
   RUNG wire#powerrail
      "LDH100_DB_1"(AI_Temp_RAW := "LDH_Temp_1", cycleTime_ms := #OB1_PREV_CYCLE, AI_Hum_RAW := "LDH_Feucht_1", Quittieren := "HMI_313".Quittieren313, Temp_filt => "Re3", Hum_filt => "Re4", Temp_real => "Re1", Hum_real => "Re2", Warnung => "B1", OK => "B2", SensorError_Temp => "B3", SensorError_Hum => "B4", SensorDefekt => "B5", Strom_Hum_mA => "Re6", Strom_Temp_mA => "Re5", Alarm_Temp => "B6", Alarm_Hum => "B7")
   END_RUNG
   // the same network as SCL:
   "LDH100_DB_1"(AI_Temp_RAW := "LDH_Temp_1",   // "LDH100"
                 cycleTime_ms := #OB1_PREV_CYCLE,
                 AI_Hum_RAW := "LDH_Feucht_1",
                 Quittieren := "HMI_313".Quittieren313,
                 Temp_filt => "Re3",
                 Hum_filt => "Re4",
                 Temp_real => "Re1",
                 Hum_real => "Re2",
                 Warnung => "B1",
                 OK => "B2",
                 SensorError_Temp => "B3",
                 SensorError_Hum => "B4",
                 SensorDefekt => "B5",
                 Strom_Hum_mA => "Re6",
                 Strom_Temp_mA => "Re5",
                 Alarm_Temp => "B6",
                 Alarm_Hum => "B7");
END_REGION

REGION Network 2
   RUNG wire#powerrail
      "LDH100_DB_2"(AI_Temp_RAW := "LDH_Temp_2", cycleTime_ms := #OB1_PREV_CYCLE, AI_Hum_RAW := "LDH_Feucht_2", Quittieren := "HMI_313".Quittieren313, Temp_filt =>, Hum_filt =>, Temp_real =>, Hum_real =>, Warnung =>, OK =>, SensorError_Temp =>, SensorError_Hum =>, SensorDefekt =>, Strom_Hum_mA =>, Strom_Temp_mA =>, Alarm_Temp =>, Alarm_Hum =>)
   END_RUNG
   // the same network as SCL:
   "LDH100_DB_2"(AI_Temp_RAW := "LDH_Temp_2",   // "LDH100"
                 cycleTime_ms := #OB1_PREV_CYCLE,
                 AI_Hum_RAW := "LDH_Feucht_2",
                 Quittieren := "HMI_313".Quittieren313);
END_REGION

REGION Network 3
   RUNG wire#powerrail
      "GILL4212_DB"(AI_Fine_RAW := "Gill_Fine", AI_Coarse_RAW := "Gill_Coarse", AI_Water_RAW := "Gill_Water", Quittieren := "HMI_313".Quittieren313, Fine_percent =>, Coarse_percent =>, Water_percent =>, Alarm_Wear =>, Alarm_Water =>, Warnung =>, SensorError_Coarse =>, SensorError_Water =>, SensorError_Fine =>, OK =>)
   END_RUNG
   // the same network as SCL:
   "GILL4212_DB"(AI_Fine_RAW := "Gill_Fine",   // "GILL4212"
                 AI_Coarse_RAW := "Gill_Coarse",
                 AI_Water_RAW := "Gill_Water",
                 Quittieren := "HMI_313".Quittieren313);
END_REGION

REGION Network 4
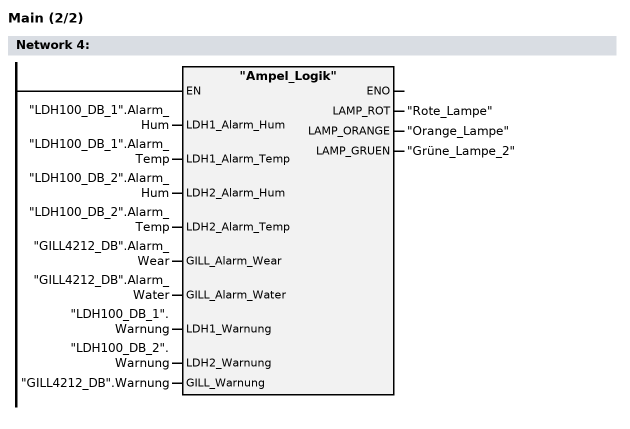
   RUNG wire#powerrail
      "Ampel_Logik"(LDH1_Alarm_Hum := "LDH100_DB_1".Alarm_Hum, LDH1_Alarm_Temp := "LDH100_DB_1".Alarm_Temp, LDH2_Alarm_Hum := "LDH100_DB_2".Alarm_Hum, LDH2_Alarm_Temp := "LDH100_DB_2".Alarm_Temp, GILL_Alarm_Wear := "GILL4212_DB".Alarm_Wear, GILL_Alarm_Water := "GILL4212_DB".Alarm_Water, LDH1_Warnung := "LDH100_DB_1".Warnung, LDH2_Warnung := "LDH100_DB_2".Warnung, GILL_Warnung := "GILL4212_DB".Warnung, LAMP_ROT => "Rote_Lampe", LAMP_ORANGE => "Orange_Lampe", LAMP_GRUEN => "Grüne_Lampe_2")
   END_RUNG
   // the same network as SCL:
   "Ampel_Logik"(LDH1_Alarm_Hum := "LDH100_DB_1".Alarm_Hum,
                 LDH1_Alarm_Temp := "LDH100_DB_1".Alarm_Temp,
                 LDH2_Alarm_Hum := "LDH100_DB_2".Alarm_Hum,
                 LDH2_Alarm_Temp := "LDH100_DB_2".Alarm_Temp,
                 GILL_Alarm_Wear := "GILL4212_DB".Alarm_Wear,
                 GILL_Alarm_Water := "GILL4212_DB".Alarm_Water,
                 LDH1_Warnung := "LDH100_DB_1".Warnung,
                 LDH2_Warnung := "LDH100_DB_2".Warnung,
                 GILL_Warnung := "GILL4212_DB".Warnung,
                 LAMP_ROT => "Rote_Lampe",
                 LAMP_ORANGE => "Orange_Lampe",
                 LAMP_GRUEN => "Grüne_Lampe_2");
END_REGION
END_ORGANIZATION_BLOCK

(* ===== HMI "HMI_RT" =====
system functions are stored by id; their names below are inferred from use
connection "HMI_Verbindung_1": IF1 B, SIMATIC S7 300/400 MPI
connection "HMI_Verbindung_3": ETHERNET, S7_1500_OMS

HMI tags "_test"
   "LDH100_DB_1_Temp_real" : Real = PLC LDH100_DB_1.Temp_real AT %DB1.DBD16, 1 s
   "LDH100_DB_1_Temp_filt" : Real = PLC LDH100_DB_1.Temp_filt AT %DB1.DBD8, 1 s
   "LDH100_DB_1_TempGrenze_Alarm" : Real = PLC LDH100_DB_1.TempGrenze_Alarm AT %DB1.DBD38, 1 s
   "LDH100_DB_1_Strom_Temp_mA" : Real = PLC LDH100_DB_1.Strom_Temp_mA AT %DB1.DBD30, 1 s
   "LDH100_DB_1_Hum_real" : Real = PLC LDH100_DB_1.Hum_real AT %DB1.DBD20, 1 s
   "LDH100_DB_1_Hum_filt" : Real = PLC LDH100_DB_1.Hum_filt AT %DB1.DBD12, 1 s
   "LDH100_DB_1_HumGrenze_Alarm" : Real = PLC LDH100_DB_1.HumGrenze_Alarm AT %DB1.DBD42, 1 s
   "LDH100_DB_1_Strom_Hum_mA" : Real = PLC LDH100_DB_1.Strom_Hum_mA AT %DB1.DBD26, 1 s
   "GILL4212_DB_Fine_percent" : Real = PLC GILL4212_DB.Fine_percent AT %DB3.DBD8, 1 s
   "GILL4212_DB_Coarse_percent" : Real = PLC GILL4212_DB.Coarse_percent AT %DB3.DBD12, 1 s
   "GILL4212_DB_Water_percent" : Real = PLC GILL4212_DB.Water_percent AT %DB3.DBD16, 1 s
   "LDH100_DB_2_Temp_real" : Real = PLC LDH100_DB_2.Temp_real AT %DB2.DBD16, 1 s
   "LDH100_DB_2_Temp_filt" : Real = PLC LDH100_DB_2.Temp_filt AT %DB2.DBD8, 1 s
   "LDH100_DB_2_TempGrenze_Alarm" : Real = PLC LDH100_DB_2.TempGrenze_Alarm AT %DB2.DBD38, 1 s
   "LDH100_DB_2_Strom_Temp_mA" : Real = PLC LDH100_DB_2.Strom_Temp_mA AT %DB2.DBD30, 1 s
   "LDH100_DB_2_Hum_real" : Real = PLC LDH100_DB_2.Hum_real AT %DB2.DBD20, 1 s
   "LDH100_DB_2_Hum_filt" : Real = PLC LDH100_DB_2.Hum_filt AT %DB2.DBD12, 1 s
   "LDH100_DB_2_HumGrenze_Alarm" : Real = PLC LDH100_DB_2.HumGrenze_Alarm AT %DB2.DBD42, 1 s
   "LDH100_DB_2_Strom_Hum_mA" : Real = PLC LDH100_DB_2.Strom_Hum_mA AT %DB2.DBD26, 1 s
   "Grüne_Lampe_2" : Bool = PLC Grüne_Lampe_2 AT %I124.2, 1 s
   "Orange_Lampe" : Bool = PLC Orange_Lampe AT %I124.1, 1 s
   "Rote_Lampe" : Bool = PLC Rote_Lampe AT %I124.0, 1 s
   "HMI_313_Quittieren313" : Bool = PLC HMI_313.Quittieren313 AT %DB4.DBX0.0, 1 s
   "LDH100_DB_1_Temp_real(1)" : Real = PLC LDH100_DB_1.Temp_real, 1 s
   "LDH100_DB_1_Temp_filt(1)" : Real = PLC LDH100_DB_1.Temp_filt, 1 s
   "LDH100_DB_1_TempGrenze_Alarm(1)" : Real = PLC LDH100_DB_1.TempGrenze_Alarm, 1 s
   "LDH100_DB_1_Strom_Temp_mA(1)" : Real = PLC LDH100_DB_1.Strom_Temp_mA, 1 s
   "GILL4212_DB_Fine_percent(1)" : Real = PLC GILL4212_DB.Fine_percent, 1 s
   "GILL4212_DB_Coarse_percent(1)" : Real = PLC GILL4212_DB.Coarse_percent, 1 s
   "GILL4212_DB_Water_percent(1)" : Real = PLC GILL4212_DB.Water_percent, 1 s
   "LDH100_DB_2_Temp_real(1)" : Real = PLC LDH100_DB_2.Temp_real, 1 s
   "LDH100_DB_2_TempGrenze_Alarm(1)" : Real = PLC LDH100_DB_2.TempGrenze_Alarm, 1 s
   "LDH100_DB_2_Strom_Temp_mA(1)" : Real = PLC LDH100_DB_2.Strom_Temp_mA, 1 s
   "LDH100_DB_2_Hum_real(1)" : Real = PLC LDH100_DB_2.Hum_real, 1 s
   "LDH100_DB_1_Hum_real(1)" : Real = PLC LDH100_DB_1.Hum_real, 1 s
   "LDH100_DB_1_Hum_filt(1)" : Real = PLC LDH100_DB_1.Hum_filt, 1 s
   "Grüne_Lampe_2(1)" : Bool = PLC "Grüne_Lampe_2(1)" AT %Q0.2, 1 s
   "Orange_Lampe(1)" : Bool = PLC "Orange_Lampe(1)" AT %Q0.1, 1 s
   "Rote_Lampe(1)" : Bool = PLC "Rote_Lampe(1)" AT %Q0.0, 1 s
   "HMI_Quittieren1500" : Bool = PLC HMI.Quittieren1500, 1 s
   "LDH100_DB_1_Strom_Hum_mA(1)" : Real = PLC LDH100_DB_1.Strom_Hum_mA, 1 s
   "LDH100_DB_2_Strom_Hum_mA(1)" : Real = PLC LDH100_DB_2.Strom_Hum_mA, 1 s
   "LDH100_DB_1_HumGrenze_Alarm(1)" : Real = PLC LDH100_DB_1.HumGrenze_Alarm, 1 s

HMI tags "Variablentabelle_1"
   "Quittierung" : Bool, internal

screen "Messwerte313" 1920x1080
   GraphicView "Grafikanzeige_1" at 1240,60 size 504x176; Picture "ChatGPT Image 26. Mai 2025, 09_14_11"
   Circle "Kreis_1" at 1135,977 size 75x75
      Appearance <- "Grüne_Lampe_2"
   Circle "Kreis_2" at 1234,977 size 75x75
      Appearance <- "Orange_Lampe"
   Circle "Kreis_3" at 1339,977 size 75x75
      Appearance <- "Rote_Lampe"
   Button "Schaltfläche_1" at 1493,987 size 205x56; TextOff 'Quittieren'
      on Press: function_b14e0dd5("HMI_313_Quittieren313", 0)
   IOField "EA-Feld_1" at 84,165 size 152x49; FormatPattern s99.9; Unit  °C
      ProcessValue <- "LDH100_DB_1_Temp_real"
   IOField "EA-Feld_2" at 245,165 size 135x49; FormatPattern 99.9; Unit  %
      ProcessValue <- "LDH100_DB_1_Hum_real"
   IOField "EA-Feld_3" at 82,268 size 134x49; FormatPattern 99.9; Unit  °C
      ProcessValue <- "LDH100_DB_1_TempGrenze_Alarm"
   IOField "EA-Feld_4" at 247,268 size 135x49; FormatPattern 99.9; Unit  %
      ProcessValue <- "LDH100_DB_1_HumGrenze_Alarm"
   TextField "Textfeld_5" at 86,114 size 429x39; Text 'Getriebekammer'
   IOField "EA-Feld_5" at 451,269 size 134x49; FormatPattern 99.9; Unit  °C
      ProcessValue <- "LDH100_DB_2_TempGrenze_Alarm"
   IOField "EA-Feld_6" at 609,269 size 135x49; FormatPattern 99.9; Unit  %
      ProcessValue <- "LDH100_DB_2_HumGrenze_Alarm"
   TextField "Textfeld_8" at 452,116 size 547x39; Text 'Emulsionkammer'
   IOField "EA-Feld_7" at 451,166 size 152x49; FormatPattern s99.9; Unit  °C
      ProcessValue <- "LDH100_DB_2_Temp_real"
   IOField "EA-Feld_8" at 609,165 size 135x49; FormatPattern 99.9; Unit  %
      ProcessValue <- "LDH100_DB_2_Hum_real"
   TextField "Textfeld_11" at 855,1005 size 365x39; Text 'Zustand'
   Bar "Balken_1" at 78,463 size 278x117; MinimumValue 0; MaximumValue 100
      ProcessValue <- "GILL4212_DB_Fine_percent"
   Bar "Balken_2" at 448,464 size 278x117; MinimumValue 0; MaximumValue 100
      ProcessValue <- "GILL4212_DB_Coarse_percent"
   TextField "Textfeld_12" at 77,422 size 102x39; Text 'Fine'
   TextField "Textfeld_13" at 448,423 size 139x39; Text 'Coarse'
   TextField "Textfeld_14" at 58,368 size 570x43; Text 'Verschleiss'
   Bar "Balken_3" at 76,650 size 278x117; MinimumValue 0; MaximumValue 100
      ProcessValue <- "GILL4212_DB_Water_percent"
   TextField "Textfeld_1" at 69,603 size 415x39; Text 'Wasserkontamination'
   TrendView "Kurvenanzeige_1" at 860,250 size 963x602
   IOField "EA-Feld_9" at 247,318 size 125x35; FormatPattern 99.999; Unit  mA
      ProcessValue <- "LDH100_DB_1_Strom_Hum_mA"
   IOField "EA-Feld_10" at 82,318 size 125x35; FormatPattern 99.999; Unit  mA
      ProcessValue <- "LDH100_DB_1_Strom_Temp_mA"
   IOField "EA-Feld_11" at 451,318 size 125x35; FormatPattern 99.999; Unit  mA
      ProcessValue <- "LDH100_DB_2_Strom_Temp_mA"
   IOField "EA-Feld_12" at 610,318 size 125x35; FormatPattern 99.999; Unit  mA
      ProcessValue <- "LDH100_DB_2_Strom_Hum_mA"
   IOField "EA-Feld_13" at 84,214 size 152x49; FormatPattern s99.9; Unit  °C
      ProcessValue <- "LDH100_DB_1_Temp_filt"
   IOField "EA-Feld_14" at 245,214 size 152x49; FormatPattern s99.9; Unit  °C
      ProcessValue <- "LDH100_DB_1_Hum_filt"
   IOField "EA-Feld_15" at 451,215 size 152x49; FormatPattern s99.9; Unit  °C
      ProcessValue <- "LDH100_DB_2_Temp_filt"
   IOField "EA-Feld_16" at 609,213 size 152x49; FormatPattern s99.9; Unit  °C
      ProcessValue <- "LDH100_DB_2_Hum_filt"
   TextField "Textfeld_2" at 16,171 size 66x25; Text 'IST'
   TextField "Textfeld_3" at 2,224 size 114x25; Text 'Gefiltert'
   TextField "Textfeld_4" at 5,276 size 94x25; Text 'Grenze'
   TextField "Textfeld_6" at 21,21 size 189x39; Text 'S7-300 Test'
   Softkey "[!Invalid!]Softkey_F2" at 0,0 size 0x0
      on KeyDown: ActivateScreen("Messwerte1500", 0)
   Softkey "[!Invalid!]Softkey_F1" at 0,0 size 0x0
      on KeyDown: ActivateScreen("Messwerte313", 0)

screen "Messwerte1500" 1920x1080
   Softkey "[!Invalid!]Softkey_F2" at 0,0 size 0x0
      on KeyDown: ActivateScreen("Messwerte1500", 0)
   Softkey "[!Invalid!]Softkey_F1" at 0,0 size 0x0
      on KeyDown: ActivateScreen("Messwerte313", 0)
   GraphicView "Grafikanzeige_1" at 1240,60 size 504x176; Picture "ChatGPT Image 26. Mai 2025, 09_14_11"
   Circle "Kreis_1" at 1135,977 size 75x75
      Appearance <- "Grüne_Lampe_2(1)"
   Circle "Kreis_2" at 1234,977 size 75x75
      Appearance <- "Orange_Lampe(1)"
   Circle "Kreis_3" at 1339,977 size 75x75
      Appearance <- "Rote_Lampe(1)"
   Button "Schaltfläche_1" at 1493,987 size 205x56; TextOff 'Quittieren'
      on Press: function_b14e0dd5("HMI_Quittieren1500", 0)
   IOField "EA-Feld_1" at 84,165 size 152x49; FormatPattern s99.9; Unit  °C
      ProcessValue <- "LDH100_DB_1_Temp_real(1)"
   IOField "EA-Feld_2" at 245,165 size 153x49; FormatPattern s99.9; Unit  %
      ProcessValue <- "LDH100_DB_1_Hum_real(1)"
   IOField "EA-Feld_3" at 82,268 size 134x49; FormatPattern 99.9; Unit  °C
      ProcessValue <- "LDH100_DB_1_TempGrenze_Alarm(1)"
   IOField "EA-Feld_4" at 247,268 size 135x49; FormatPattern 99.9; Unit  %
      ProcessValue <- "LDH100_DB_1_HumGrenze_Alarm(1)"
   TextField "Textfeld_5" at 86,114 size 429x39; Text 'Getriebekammer'
   IOField "EA-Feld_5" at 451,269 size 134x49; FormatPattern 99.9; Unit  °C
      ProcessValue <- "LDH100_DB_2_TempGrenze_Alarm(1)"
   IOField "EA-Feld_6" at 609,269 size 135x49; FormatPattern 99.9; Unit  %
      ProcessValue <- "LDH100_DB_2_HumGrenze_Alarm"
   TextField "Textfeld_8" at 452,116 size 547x39; Text 'Emulsionkammer'
   IOField "EA-Feld_7" at 451,166 size 152x49; FormatPattern s99.9; Unit  °C
      ProcessValue <- "LDH100_DB_2_Temp_real(1)"
   IOField "EA-Feld_8" at 609,165 size 135x49; FormatPattern 99.9; Unit  %
      ProcessValue <- "LDH100_DB_2_Hum_real(1)"
   TextField "Textfeld_11" at 855,1005 size 365x39; Text 'Zustand'
   Bar "Balken_1" at 78,463 size 278x117; MinimumValue 0; MaximumValue 100
      ProcessValue <- "GILL4212_DB_Fine_percent(1)"
   Bar "Balken_2" at 448,464 size 278x117; MinimumValue 0; MaximumValue 100
      ProcessValue <- "GILL4212_DB_Coarse_percent(1)"
   TextField "Textfeld_12" at 77,422 size 102x39; Text 'Fine'
   TextField "Textfeld_13" at 448,423 size 139x39; Text 'Coarse'
   TextField "Textfeld_14" at 49,374 size 570x43; Text 'Verschleiss'
   Bar "Balken_3" at 76,650 size 278x117; MinimumValue 0; MaximumValue 100
      ProcessValue <- "GILL4212_DB_Water_percent(1)"
   TextField "Textfeld_1" at 69,603 size 415x39; Text 'Wasserkontamination'
   TrendView "Kurvenanzeige_1" at 860,250 size 963x602
   IOField "EA-Feld_9" at 248,318 size 125x35; FormatPattern 99.999; Unit  mA
      ProcessValue <- "LDH100_DB_1_Strom_Hum_mA(1)"
   IOField "EA-Feld_10" at 82,318 size 125x35; FormatPattern 99.999; Unit  mA
      ProcessValue <- "LDH100_DB_1_Strom_Temp_mA(1)"
   IOField "EA-Feld_11" at 451,318 size 125x35; FormatPattern 99.999; Unit  mA
      ProcessValue <- "LDH100_DB_2_Strom_Temp_mA(1)"
   IOField "EA-Feld_12" at 609,318 size 125x35; FormatPattern 99.999; Unit  mA
      ProcessValue <- "LDH100_DB_2_Strom_Hum_mA(1)"
   IOField "EA-Feld_13" at 84,214 size 152x49; FormatPattern s99.9; Unit  °C
      ProcessValue <- "LDH100_DB_1_Temp_filt(1)"
   IOField "EA-Feld_14" at 246,214 size 152x49; FormatPattern s99.9; Unit  °C
      ProcessValue <- "LDH100_DB_1_Hum_filt"
   IOField "EA-Feld_15" at 451,215 size 152x49; FormatPattern s99.9; Unit  °C
      ProcessValue <- "LDH100_DB_1_Temp_filt(1)"
   IOField "EA-Feld_16" at 609,214 size 152x49; FormatPattern s99.9; Unit  °C
      ProcessValue <- "LDH100_DB_1_Hum_filt(1)"
   TextField "Textfeld_2" at 7,183 size 198x25; Text 'IST'
   TextField "Textfeld_3" at 4,227 size 228x25; Text 'Gefiltert'
   TextField "Textfeld_4" at 7,279 size 184x25; Text 'Grenze'
   TextField "Textfeld_6" at 21,21 size 208x39; Text 'S7-1500 Test'
*)